Flt - Depress Man Weld To Continue FB1[301].22'; 9655 '~S001R08CN.I.Wc2SGunFlt - Weld Controller 2 Servo Gun Fault FB1[301].23'; 9656 '~S001R08CN.I.Wc2SGunMtrTempFlt - Cntrl 2 Servo Gun Motor Over Temp FB1[301].24'; 9657 '~S001R08CN.I.Td2MtrFlt - Tip Dress 2 Motor Fault FB1[301].25'; 9658 '~S001R08CN.I.WC2XfmrTempFlt - Weld Cntrl 2 Transformer Over Temp FB1[301].26'; 9659 '~S001R08CN.I.AutoTipChng2Flt - Auto Tip Changer 2 Fault FB1[301].27'; 9660 '~S001R08CN.I.Slr2NotReady - Seal Controller 2 Not Ready FB1[301].28'; 9661 '~S001R08CN.I.Slr2MajorFlt - Seal Controller 2 Major Fault FB1[301].29'; 9662 '~S001R08CN.I.Slr2VolNotOk - Seal Controller 2 Volume Not Ok Fault FB1[301].30'; 9663 '~S001R08CN.I.Slr2PurgeFlt - Seal Controller 2 Purge Fault FB1[301].31'; 9664 '~S001R08CN.I.Slr2DoserNot Filled - Seal Cntrl 2 Doser Not Filled FB1[302].0'; 9665 '~S001R08CN.I.Slr2No2ClnMxr - Seal Cntrl2 No 2C In Mixer Fault FB1[302].1'; 9666 '~S001R08CN.I.Slr2NzlBroken - Seal Controller 2 Nozzle Broken Fault FB1[302].2'; 9667 '~S001R08CN.I.Slr2NozzleChgReq - Seal Cntrl2 Nozzle Change Reqd FB1[302].3'; 9668 '~S001R08CN.I.Slr2CycleInterrupted - Seal Cntrl2 Cycle Interrupted FB1[302].4'; 9669 '~S001R08CN.I.Stdw2Flt - Stud Weld 2 Weld Fault FB1[302].5'; 9670 '~S001R08CN.I.Stdw2DlyExcdd - Stud Weld 2 Time Delay Exceeded Flt FB1[302].6'; 9671 '~S001R08CN.I.Stdw2Maint Reqd - Stud Weld 2 Maintenance Required FB1[302].7'; 9672 '~S001R08CN.I.Stdw2Reject - Stud Weld 2 art Reject Fault FB1[302].8'; 9673 '~S001R08CN.I.Rvt2Flt - Rivet Controller 2 Fault FB1[302].9'; 9674 '~S001R08CN.I.Rvt2DlyExcdd - Rivet Cntrl 2 Time Delay Exceeded Flt FB1[302].10'; 9675 '~S001R08CN.I.AutoPulledTipByp2 - Auto Pulled Tip Bypass 2 FB1[302].11'; 9676 '~S001R08CN.I.StdWld2EquipmentFlt - Stud Weld 2 Equipment Fault FB1[302].12'; 9677 '~S001R08CN.I.StdWld2BrcktNotPresent - Stud Weld 2 Bracket Not Pres FB1[302].13'; 9678 '~S001R08CN.Ix.LsrWldMntrFlt - Seam Geometry/Laser Weld Monitor Flt FB1[302].14'; 9679 '~S001R08CN.Ix.LsrHeadFlt - Laser Head Fault FB1[302].15'; 9680 '~S001R08CN.Ix.LsrGlsFlt - Glass Fault FB1[302].16'; 9681 '~S001R08CN.Ix.LsrWhlFlt - Pressure Wheel Not In Range Fault FB1[302].17'; 9682 '~S001R08CN.Ix.LsrGeoFlt - Seam Geometry/Laser Bad Process Geo Flt FB1[302].18'; 9683 '~S001R08CN.Ix.LsrHdCollFlt - Laser Head Collision Fault FB1[302].19'; 9684 '~S001R08CN.Ix.LsrHdSysFlt - Laser Head System Fault FB1[302].20'; 9685 '~S001R08CN.Ix.LsrHdFar - Laser Head Far Fault FB1[302].21'; 9686 '~S001R08CN.Ix.LsrHdSftCollFlt - Laser Head Software Collision Flt FB1[302].22'; 9687 '~S001R08CN.I.O.TipChngReqd2 - Weld Cntrl 2 Tip Change Required FB1[302].23'; 9688 '~S001R08CN.I.M.NutDetectFlt2 - Nut Welder 2 Nut Detection Fault FB1[302].24'; 9689 '~S001R08CN.I.M.NutProjFlt2 - Nut Welder 2 Weld Not In Tolerance FB1[302].25'; 9690 '~S001R08CN.I.TCWrongToolInStand - Tool Changer Wrong Tool In Stand FB1[302].26'; 9691 '~Spare FB1[302].27'; 9692 '~Spare FB1[302].28'; 9693 '~Spare FB1[302].29'; 9694 '~Spare FB1[302].30'; 9695 '~Spare FB1[302].31'; 9696 '~S001R08CN.I.VisionCommOK - Vision System Comm Fault FB1[303].0'; 9697 '~S001R08CN.I.OutOfTolerance - Vision System Out Of Tolerance FB1[303].1'; 9698 '~S001R08CN.I.MeasureReject - Vision System Measure Reject FB1[303].2'; 9699 '~S001R08CN.I.VisionSysCalibrationFlt - Vision System Calibration Flt FB1[303].3'; 9700 '~S001R08CN.I.VisionSysFlt - Vision System Flt FB1[303].4'; 9701 '~Spare FB1[303].5'; 9702 '~Spare FB1[303].6'; 9703 '~Spare FB1[303].7'; 9704 '~Spare FB1[303].8'; 9705 '~Spare FB1[303].9'; 9706 '~Spare FB1[303].10'; 9707 '~Spare FB1[303].11'; 9708 '~Spare FB1[303].12'; 9709 '~Spare FB1[303].13'; 9710 '~Spare FB1[303].14'; 9711 '~Spare FB1[303].15'; 9712 '~Spare FB1[303].16'; 9713 '~Spare FB1[303].17'; 9714 '~S001R08CN.M.InteruptCyc - Laser Cyc Interupt Cut Wire And Reject Car FB1[303].18'; 9715 '~S001R08CN.M.SuspectPart Inspect Vehicle And Accept Or Reject FB1[303].19'; 9716 '~S001R08 Power Meter High Power Fault Detected FB1[303].20'; 9717 '~S001R08 Power Meter Low Power Fault Detected FB1[303].21'; 9718 '~Spare FB1[303].22'; 9719 '~Spare FB1[303].23'; 9720 '~Spare FB1[303].24'; 9721 '~Spare FB1[303].25'; 9722 '~Spare FB1[303].26'; 9723 '~Spare FB1[303].27'; 9724 '~Spare FB1[303].28'; 9725 '~Spare FB1[303].29'; 9726 '~Spare FB1[303].30'; 9727 '~Spare FB1[303].31'; 9728 '~Spare FB1[304].0'; 9729 '~Spare FB1[304].1'; 9730 '~Spare FB1[304].2'; 9731 '~Spare FB1[304].3'; 9732 '~Spare FB1[304].4'; 9733 '~Spare FB1[304].5'; 9734 '~Spare FB1[304].6'; 9735 '~Spare FB1[304].7'; 9736 '~Spare FB1[304].8'; 9737 '~Spare FB1[304].9'; 9738 '~Spare FB1[304].10'; 9739 '~Spare FB1[304].11'; 9740 '~Spare FB1[304].12'; 9741 '~Spare FB1[304].13'; 9742 '~Spare FB1[304].14'; 9743 '~Spare FB1[304].15'; 9744 '~Spare FB1[304].16'; 9745 '~Spare FB1[304].17'; 9746 '~Spare FB1[304].18'; 9747 '~Spare FB1[304].19'; 9748 '~Spare FB1[304].20'; 9749 '~Spare FB1[304].21'; 9750 '~Spare FB1[304].22'; 9751 '~Spare FB1[304].23'; 9752 '~Spare FB1[304].24'; 9753 '~Spare FB1[304].25'; 9754 '~Spare FB1[304].26'; 9755 '~Spare FB1[304].27'; 9756 '~Spare FB1[304].28'; 9757 '~Spare FB1[304].29'; 9758 '~Spare FB1[304].30'; 9759 '~Spare FB1[304].31'; 9760 '~Spare FB1[305].0'; 9761 '~Spare FB1[305].1'; 9762 '~Spare FB1[305].2'; 9763 '~Spare FB1[305].3'; 9764 '~Spare FB1[305].4'; 9765 '~Spare FB1[305].5'; 9766 '~Spare FB1[305].6'; 9767 '~Spare FB1[305].7'; 9768 '~Spare FB1[305].8'; 9769 '~Spare FB1[305].9'; 9770 '~Spare FB1[305].10'; 9771 '~Spare FB1[305].11'; 9772 '~Spare FB1[305].12'; 9773 '~Spare FB1[305].13'; 9774 '~Spare FB1[305].14'; 9775 '~Spare FB1[305].15'; 9776 '~Spare FB1[305].16'; 9777 '~Spare FB1[305].17'; 9778 '~Spare FB1[305].18'; 9779 '~Spare FB1[305].19'; 9780 '~Spare FB1[305].20'; 9781 '~Spare FB1[305].21'; 9782 '~Spare FB1[305].22'; 9783 '~Spare FB1[305].23'; 9784 '~Spare FB1[305].24'; 9785 '~Spare FB1[305].25'; 9786 '~Spare FB1[305].26'; 9787 '~Spare FB1[305].27'; 9788 '~Spare FB1[305].28'; 9789 '~Spare FB1[305].29'; 9790 '~Spare FB1[305].30'; 9791 '~Spare FB1[305].31'; 9792 '~Spare FB1[306].0'; 9793 '~Spare FB1[306].1'; 9794 '~Spare FB1[306].2'; 9795 '~Spare FB1[306].3'; 9796 '~Spare FB1[306].4'; 9797 '~Spare FB1[306].5'; 9798 '~Spare FB1[306].6'; 9799 '~Spare FB1[306].7'; 9800 '~Spare FB1[306].8'; 9801 '~Spare FB1[306].9'; 9802 '~Spare FB1[306].10'; 9803 '~Spare FB1[306].11'; 9804 '~Spare FB1[306].12'; 9805 '~Spare FB1[306].13'; 9806 '~Spare FB1[306].14'; 9807 '~Spare FB1[306].15'; 9808 '~Spare FB1[306].16'; 9809 '~Spare FB1[306].17'; 9810 '~Spare FB1[306].18'; 9811 '~Spare FB1[306].19'; 9812 '~Spare FB1[306].20'; 9813 '~Spare FB1[306].21'; 9814 '~Spare FB1[306].22'; 9815 '~Spare FB1[306].23'; 9816 '~Spare FB1[306].24'; 9817 '~Spare FB1[306].25'; 9818 '~Spare FB1[306].26'; 9819 '~Spare FB1[306].27'; 9820 '~Spare FB1[306].28'; 9821 '~Spare FB1[306].29'; 9822 '~Spare FB1[306].30'; 9823 '~Spare FB1[306].31'; 9824 '~Spare FB1[307].0'; 9825 '~Spare FB1[307].1'; 9826 '~Spare FB1[307].2'; 9827 '~Spare FB1[307].3'; 9828 '~Spare FB1[307].4'; 9829 '~Spare FB1[307].5'; 9830 '~Spare FB1[307].6'; 9831 '~Spare FB1[307].7'; 9832 '~Spare FB1[307].8'; 9833 '~Spare FB1[307].9'; 9834 '~Spare FB1[307].10'; 9835 '~Spare FB1[307].11'; 9836 '~Spare FB1[307].12'; 9837 '~Spare FB1[307].13'; 9838 '~Spare FB1[307].14'; 9839 '~Spare FB1[307].15'; 9840 '~Spare FB1[307].16'; 9841 '~Spare FB1[307].17'; 9842 '~Spare FB1[307].18'; 9843 '~Spare FB1[307].19'; 9844 '~Spare FB1[307].20'; 9845 '~Spare FB1[307].21'; 9846 '~Spare FB1[307].22'; 9847 '~Spare FB1[307].23'; 9848 '~Spare FB1[307].24'; 9849 '~Spare FB1[307].25'; 9850 '~Spare FB1[307].26'; 9851 '~Spare FB1[307].27'; 9852 '~Spare FB1[307].28'; 9853 '~Spare FB1[307].29'; 9854 '~Spare FB1[307].30'; 9855 '~Spare FB1[307].31'; 9856 '~Spare FB1[308].0'; 9857 '~Spare FB1[308].1'; 9858 '~Spare FB1[308].2'; 9859 '~Spare FB1[308].3'; 9860 '~Spare FB1[308].4'; 9861 '~Spare FB1[308].5'; 9862 '~Spare FB1[308].6'; 9863 '~Spare FB1[308].7'; 9864 '~Spare FB1[308].8'; 9865 '~Spare FB1[308].9'; 9866 '~Spare FB1[308].10'; 9867 '~Spare FB1[308].11'; 9868 '~Spare FB1[308].12'; 9869 '~Spare FB1[308].13'; 9870 '~Spare FB1[308].14'; 9871 '~Spare FB1[308].15'; 9872 '~Spare FB1[308].16'; 9873 '~Spare FB1[308].17'; 9874 '~Spare FB1[308].18'; 9875 '~Spare FB1[308].19'; 9876 '~Spare FB1[308].20'; 9877 '~Spare FB1[308].21'; 9878 '~Spare FB1[308].22'; 9879 '~Spare FB1[308].23'; 9880 '~Spare FB1[308].24'; 9881 '~Spare FB1[308].25'; 9882 '~Spare FB1[308].26'; 9883 '~Spare FB1[308].27'; 9884 '~Spare FB1[308].28'; 9885 '~Spare FB1[308].29'; 9886 '~Spare FB1[308].30'; 9887 '~Spare FB1[308].31'; 9888 '~Spare FB1[309].0'; 9889 '~Spare FB1[309].1'; 9890 '~Spare FB1[309].2'; 9891 '~Spare FB1[309].3'; 9892 '~Spare FB1[309].4'; 9893 '~Spare FB1[309].5'; 9894 '~Spare FB1[309].6'; 9895 '~Spare FB1[309].7'; 9896 '~Spare FB1[309].8'; 9897 '~Spare FB1[309].9'; 9898 '~Spare FB1[309].10'; 9899 '~Spare FB1[309].11'; 9900 '~Spare FB1[309].12'; 9901 '~Spare FB1[309].13'; 9902 '~Spare FB1[309].14'; 9903 '~Spare FB1[309].15'; 9904 '~Spare FB1[309].16'; 9905 '~Spare FB1[309].17'; 9906 '~Spare FB1[309].18'; 9907 '~Spare FB1[309].19'; 9908 '~Spare FB1[309].20'; 9909 '~Spare FB1[309].21'; 9910 '~Spare FB1[309].22'; 9911 '~Spare FB1[309].23'; 9912 '~Spare FB1[309].24'; 9913 '~Spare FB1[309].25'; 9914 '~Spare FB1[309].26'; 9915 '~Spare FB1[309].27'; 9916 '~Spare FB1[309].28'; 9917 '~Spare FB1[309].29'; 9918 '~Spare FB1[309].30'; 9919 '~Spare FB1[309].31'; 9920 '~Spare FB1[310].0'; 9921 '~Spare FB1[310].1'; 9922 '~Spare FB1[310].2'; 9923 '~Spare FB1[310].3'; 9924 '~Spare FB1[310].4'; 9925 '~Spare FB1[310].5'; 9926 '~Spare FB1[310].6'; 9927 '~Spare FB1[310].7'; 9928 '~Spare FB1[310].8'; 9929 '~Spare FB1[310].9'; 9930 '~Spare FB1[310].10'; 9931 '~Spare FB1[310].11'; 9932 '~Spare FB1[310].12'; 9933 '~Spare FB1[310].13'; 9934 '~Spare FB1[310].14'; 9935 '~Spare FB1[310].15'; 9936 '~Spare FB1[310].16'; 9937 '~Spare FB1[310].17'; 9938 '~Spare FB1[310].18'; 9939 '~Spare FB1[310].19'; 9940 '~Spare FB1[310].20'; 9941 '~Spare FB1[310].21'; 9942 '~Spare FB1[310].22'; 9943 '~Spare FB1[310].23'; 9944 '~Spare FB1[310].24'; 9945 '~Spare FB1[310].25'; 9946 '~Spare FB1[310].26'; 9947 '~Spare FB1[310].27'; 9948 '~Spare FB1[310].28'; 9949 '~Spare FB1[310].29'; 9950 '~Spare FB1[310].30'; 9951 '~Spare FB1[310].31'; 9952 '~Spare FB1[311].0'; 9953 '~Spare FB1[311].1'; 9954 '~Spare FB1[311].2'; 9955 '~Spare FB1[311].3'; 9956 '~Spare FB1[311].4'; 9957 '~Spare FB1[311].5'; 9958 '~Spare FB1[311].6'; 9959 '~Spare FB1[311].7'; 9960 '~Spare FB1[311].8'; 9961 '~Spare FB1[311].9'; 9962 '~Spare FB1[311].10'; 9963 '~Spare FB1[311].11'; 9964 '~Spare FB1[311].12'; 9965 '~Spare FB1[311].13'; 9966 '~Spare FB1[311].14'; 9967 '~Spare FB1[311].15'; 9968 '~Spare FB1[311].16'; 9969 '~Spare FB1[311].17'; 9970 '~Spare FB1[311].18'; 9971 '~Spare FB1[311].19'; 9972 '~Spare FB1[311].20'; 9973 '~Spare FB1[311].21'; 9974 '~Spare FB1[311].22'; 9975 '~Spare FB1[311].23'; 9976 '~Spare FB1[311].24'; 9977 '~Spare FB1[311].25'; 9978 '~Spare FB1[311].26'; 9979 '~Spare FB1[311].27'; 9980 '~Spare FB1[311].28'; 9981 '~Spare FB1[311].29'; 9982 '~Spare FB1[311].30'; 9983 '~Spare FB1[311].31'; 9984 '~Spare FB1[312].0'; 9985 '~Spare FB1[312].1'; 9986 '~Spare FB1[312].2'; 9987 '~Spare FB1[312].3'; 9988 '~Spare FB1[312].4'; 9989 '~Spare FB1[312].5'; 9990 '~Spare FB1[312].6'; 9991 '~Spare FB1[312].7'; 9992 '~Spare FB1[312].8'; 9993 '~Spare FB1[312].9'; 9994 '~Spare FB1[312].10'; 9995 '~Spare FB1[312].11'; 9996 '~Spare FB1[312].12'; 9997 '~Spare FB1[312].13'; 9998 '~Spare FB1[312].14'; 9999 '~Spare FB1[312].15'; 10000 '**Local Message Display**'

text list "Text_list_IO_System": 1 'IO System 1'; 2 'IO System 2'; 3 'IO System 3'; 4 'IO System 4'

text list "G120D_Faults_Warnings": 1000 'F01000 - Internal software error'; 1001 'F01001 - FloatingPoint exception'; 1002 'F01002 - Internal software error'; 1003 'F01003 - Acknowledgment delay when accessing the memory'; 1004 'N01004 (F, A) - Internal software error'; 1005 'F01005 - File upload/download error'; 1009 'A01009 (N) - CU: Control module overtemperature'; 1010 'F01010 - Drive type unknown'; 1015 'F01015 - Internal software error'; 1016 'A01016 (F) - Firmware changed'; 1017 'A01017 - Component lists changed'; 1018 'F01018 - Booting has been interrupted several times'; 1019 'A01019 - Writing to the removable data medium unsuccessful'; 1020 'A01020 - Writing to RAM disk unsuccessful'; 1021 'A01021 - Removable data medium as USB data storage medium from the PC used'; 1023 'F01023 - Software timeout (internal)'; 1028 'A01028 (F) - Configuration error'; 1030 'F01030 - Sign-of-life failure for master control'; 1033 'F01033 - Units changeover: Reference parameter value invalid'; 1034 'F01034 - Units changeover: Calculation parameter values after reference value change unsuccessful'; 1035 'A01035 (F) - ACX: Parameter back-up file corrupted'; 1036 'F01036 (A) - ACX: Parameter back-up file missing'; 1038 'F01038 (A) - ACX: Loading the parameter back-up file unsuccessful'; 1039 'F01039 (A) - ACX: Writing to the parameter back-up file was unsuccessful'; 1040 'F01040 - Save parameter settings and carry out a POWER ON'; 1042 'F01042 - Parameter error during project download'; 1043 'F01043 - Fatal error at project download'; 1044 'F01044 - CU: Descriptive data error'; 1045 'A01045 - Configuring data invalid'; 1049 'A01049 - It is not possible to write to file'; 1054 'F01054 - CU: System limit exceeded'; 1064 'A01064 (F) - CU: Internal error (CRC)'; 1066 'A01066 - Buffer memory: 70% fill level reached or exceeded'; 1067 'A01067 - Buffer memory: 100 % fill level reached'; 1068 'F01068 - CU: Data memory memory overflow'; 1069 'A01069 - Parameter backup and device incompatible'; 1072 'F01072 - Memory card restored from the backup copy'; 1073 'A01073 (N) - POWER ON required for backup copy on memory card'; 1105 'F01105 (A) - CU: Insufficient memory'; 1107 'F01107 - Save to memory card unsuccessful'; 1112 'F01112 - CU: Power unit not permissible'; 1120 'F01120 (A) - Terminal initialization has failed'; 1122 'F01122 (A) - Frequency at the measuring probe input too high'; 1152 'F01152 - CU: Invalid constellation of drive object types'; 1205 'F01205 - CU: Time slice overflow'; 1250 'F01250 - CU: CU-EEPROM incorrect read-only data'; 1251 'A01251 - CU: CU-EEPROM incorrect read-write data'; 1257 'F01257 - CU: Firmware version out of date'; 1340 'F01340 - Topology: Too many components on one line'; 1505 'F01505 (A) - BICO: Interconnection cannot be established'; 1510 'F01510 - BICO: Signal source is not float type'; 1511 'F01511 (A) - BICO: Interconnection with different scalings'; 1512 'F01512 - BICO: No scaling available'; 1513 'F01513 (N, A) - BICO: Interconnection cross DO with different scalings'; 1514 'A01514 (F) - BICO: Error when writing during a reconnect'; 1515 'F01515 (A) - BICO: Writing to parameter not permitted as the master control is active'; 1590 'A01590 (F) - Drive: Motor maintenance interval expired'; 1600 'F01600 - SI P1 (CU): STOP A initiated'; 1611 'F01611 (A) - SI P1 (CU): Defect in a monitoring channel'; 1620 'N01620 (F, A) - SI P1 (CU): Safe Torque Off active'; 1625 'F01625 - SI P1 (CU): Sign-of-life error in safety data'; 1640 'F01640 - SI P1 (CU): component replacement identified and acknowledgment/save required'; 1641 'F01641 - SI P1 (CU): component replacement identified and save required'; 1649 'F01649 - SI P1 (CU): Internal software error'; 1650 'F01650 - SI P1 (CU): Acceptance test required'; 1651 'F01651 - SI P1 (CU): Synchronization safety time slices unsuccessful'; 1653 'F01653 - SI P1 (CU): PROFIBUS/PROFINET configuration error'; 1654 'A01654 (F) - SI P1 (CU): Deviating PROFIsafe configuration'; 1655 'F01655 - SI P1 (CU): Align monitoring functions'; 1656 'F01656 - SI P1 (CU): Parameter processor 2 error'; 1658 'F01658 - SI P1 (CU): PROFIsafe telegram number not suitable'; 1659 'F01659 - SI P1 (CU): Write request for parameter rejected'; 1660 'F01660 - SI P1 (CU): Safety-related functions not supported'; 1661 'F01661 - SI P1 (CU): Simulation of the safety inputs active'; 1662 'F01662 - Error internal communications'; 1663 'F01663 - SI P1 (CU): Copying the SI parameters rejected'; 1665 'F01665 - SI P1 (CU): System is defective'; 1666 'A01666 (F) - SI Motion P1 (CU): Steady-state (static) 1 signal at the F-DI for safe acknowledgment'; 1669 'A01669 (F, N) - SI Motion: Unfavorable combination of motor and power unit'; 1680 'F01680 - SI Motion P1 (CU): Checksum error safety monitoring functions'; 1681 'F01681 - SI Motion P1 (CU): Incorrect parameter value'; 1682 'F01682 - SI Motion P1 (CU): Monitoring function not supported'; 1683 'F01683 - SI Motion P1 (CU): SLS enable missing'; 1690 'F01690 - SI Motion: Data save problem for the NVRAM'; 1692 'F01692 - SI Motion P1 (CU): Parameter value not permitted for encoderless'; 1693 'A01693 (F) - SI P1 (CU): Safety parameter setting changed, POWER ON required'; 1696 'A01696 (F) - SI Motion: Test stop for the motion monitoring functions selected when booting'; 1697 'A01697 (F) - SI Motion: Test stop for motion monitoring functions required'; 1698 'A01698 (F) - SI P1 (CU): Commissioning mode active'; 1699 'A01699 (F) - SI P1 (CU): Test stop for STO required'; 1700 'C01700 - SI Motion P1 (CU): STOP A initiated'; 1701 'C01701 - SI Motion P1 (CU): STOP B initiated'; 1706 'C01706 - SI Motion P1 (CU): SAM/SBR limit exceeded'; 1711 'C01711 - SI Motion P1 (CU): Defect in a monitoring channel'; 1712 'C01712 - SI Motion P1 (CU): Defect in F-IO processing'; 1714 'C01714 - SI Motion P1 (CU): Safely Limited Speed exceeded'; 1716 'C01716 - SI Motion P1 (CU): Tolerance for safe motion direction exceeded'; 1770 'C01770 - SI Motion P1 (CU): Discrepancy error of the fail-safe inputs'; 1772 'A01772 - SI Motion P1 (CU): Test stop for fail-safe digital outputs running'; 1773 'F01773 - SI Motion P1 (CU): Test stop fail-safe digital output error'; 1774 'A01774 - SI Motion P1 (CU): Test stop for fail-safe digital outputs required'; 1788 'A01788 - SI: Automatic test stop waits for STO deselection via motion monitoring functions'; 1790 'A01790 - SI: Power up stopped due to STO via terminals'; 1796 'A01796 (F, N) - SI P1 (CU): Wait for communication'; 1798 'C01798 - SI Motion P1 (CU): Test stop for motion monitoring functions running'; 1799 'C01799 - SI Motion P1 (CU): Acceptance test mode active'; 1900 'A01900 (F) - PROFIBUS: Configuration telegram error'; 1910 'F01910 (N, A) - Fieldbus interface setpoint timeout'; 1920 'A01920 (F) - PROFIBUS: Interruption cyclic connection'; 1945 'A01945 - PROFIBUS: Connection to the Publisher failed'; 1946 'F01946 (A) - PROFIBUS: Connection to the Publisher aborted'; 1951 'F01951 - CU SYNC: Synchronization application clock cycle missing'; 1953 'A01953 - CU SYNC: Synchronization not completed'; 2050 'A02050 - Trace: Start not possible'; 2051 'A02051 - Trace: recording not possible as a result of know-how protection'; 2055 'A02055 - Trace: Recording time too short'; 2056 'A02056 - Trace: Recording cycle too short'; 2057 'A02057 - Trace: Time slice clock cycle invalid'; 2058 'A02058 - Trace: Time slice clock cycle for endless trace not valid'; 2059 'A02059 - Trace: Time slice clock cycle for 2 x 8 recording channels not valid'; 2060 'A02060 - Trace: Signal to be traced missing'; 2061 'A02061 - Trace: Invalid signal'; 2062 'A02062 - Trace: Invalid trigger signal'; 2063 'A02063 - Trace: Invalid data type'; 2070 'A02070 - Trace: Parameter cannot be changed'; 2075 'A02075 - Trace: Pretrigger time too long'; 2080 'F02080 - Trace: Parameterization deleted due to unit changeover'; 2095 'A02095 - MTrace 0: multiple trace cannot be activated'; 2096 'A02096 - MTrace 0: cannot be saved'; 2097 'A02097 - MTrace 1: multiple trace cannot be activated'; 2098 'A02098 - MTrace 1: cannot be saved'; 2099 'A02099 - Trace: Insufficient Control Unit memory'; 2150 'A02150 - OA: Application cannot be loaded'; 2151 'F02151 (A) - OA: Internal software error'; 2152 'F02152 (A) - OA: Insufficient memory'; 3000 'F03000 - NVRAM fault on action'; 3001 'F03001 - NVRAM checksum incorrect'; 3505 'F03505 (N, A) - Analog input wire breakage'; 3510 'A03510 (F, N) - Calibration data not plausible'; 5000 'A05000 (N) - Power unit: Overtemperature heat sink AC inverter'; 5001 'A05001 (N) - Power unit: Overtemperature depletion layer chip'; 5002 'A05002 (N) - Power unit: Air intake overtemperature'; 5004 'A05004 (N) - Power unit: Rectifier overtemperature'; 5006 'A05006 (N) - Power unit: Overtemperature thermal model'; 5065 'A05065 (F, N) - Voltage measured values not plausible'; 6310 'F06310 (A) - Supply voltage (p0210) incorrectly parameterized'; 6921 'A06921 (N) - Braking resistor phase unsymmetry'; 6922 'F06922 - Braking resistor phase failure'; 7011 'F07011 - Drive: Motor overtemperature'; 7012 'A07012 (N) - Drive: Motor temperature model 1/3 overtemperature'; 7014 'A07014 (N) - Drive: Motor temperature model configuration alarm'; 7015 'A07015 - Drive: Motor temperature sensor alarm'; 7016 'F07016 - Drive: Motor temperature sensor fault'; 7080 'F07080 - Drive: Incorrect control parameter'; 7082 'F07082 - Macro: Execution not possible'; 7083 'F07083 - Macro: ACX file not found'; 7084 'F07084 - Macro: Condition for WaitUntil not fulfilled'; 7086 'F07086 - Units changeover: Parameter limit violation due to reference value change'; 7088 'F07088 - Units changeover: Parameter limit violation due to units changeover'; 7089 'A07089 - Changing over units: Function module activation is blocked because the units have been changed over'; 7092 'A07092 - Drive: moment of inertia estimator still not ready'; 7094 'A07094 - General parameter limit violation'; 7200 'A07200 - Drive: Master control ON command present'; 7220 'F07220 (N, A) - Drive: Master control by PLC missing'; 7300 'F07300 (A) - Drive: Line contactor feedback signal missing'; 7320 'F07320 - Drive: Automatic restart interrupted'; 7321 'A07321 - Drive: Automatic restart active'; 7330 'F07330 - Flying restart: Measured search current too low'; 7331 'F07331 - Flying restart: Function not supported'; 7404 'F07404 - Drive: DC link voltage monitoring Vdc_max'; 7409 'A07409 (N) - Drive: U/f control, current limiting controller active'; 7410 'F07410 - Drive: Current controller output limited'; 7411 'F07411 - Drive: Flux setpoint not reached when building up excitation'; 7416 'A07416 - Drive: Flux controller configuration'; 7426 'F07426 (A) - Technology controller actual value limited'; 7428 'A07428 (N) - Technology controller parameterizing error'; 7435 'F07435 (N) - Drive: Setting the ramp-function generator for sensorless vector control'; 7440 'A07440 - EPOS: Jerk time is limited'; 7441 'A07441 - LR: Save the position offset of the absolute encoder adjustment'; 7442 'F07442 (A) - LR: Multiturn does not match the modulo range'; 7443 'F07443 (A) - LR: Reference point coordinate not in the permissible range'; 7450 'F07450 (A) - LR: Standstill monitoring has responded'; 7451 'F07451 (A) - LR: Position monitoring has responded'; 7452 'F07452 (A) - LR: Following error too high'; 7453 'F07453 - LR: Position actual value preprocessing error'; 7454 'A07454 - LR: Position actual value preprocessing does not have a valid encoder'; 7455 'A07455 - EPOS: Maximum velocity limited'; 7456 'A07456 - EPOS: Setpoint velocity limited'; 7457 'A07457 - EPOS: Combination of input signals illegal'; 7458 'F07458 - EPOS: Reference cam not found'; 7459 'F07459 - EPOS: No zero mark'; 7460 'F07460 - EPOS: End of reference cam not found'; 7461 'A07461 - EPOS: Reference point not set'; 7462 'A07462 - EPOS: Selected traversing block number does not exist'; 7463 'A07463 (F) - EPOS: External block change not requested in the traversing block'; 7464 'F07464 - EPOS: Traversing block is inconsistent'; 7465 'A07465 - EPOS: Traversing block does not have a subsequent block'; 7466 'A07466 - EPOS: Traversing block number assigned a multiple number of times'; 7467 'A07467 - EPOS: Traversing block has illegal task parameters'; 7468 'A07468 - EPOS: Traversing block jump destination does not exist'; 7469 'A07469 - EPOS: Traversing block < target position < software limit switch minus'; 7470 'A07470 - EPOS: Traversing block> target position > software limit switch plus'; 7471 'A07471 - EPOS: Traversing block target position outside the modulo range'; 7472 'A07472 - EPOS: Traversing block ABS_POS/ABS_NEG not possible'; 7473 'A07473 (F) - EPOS: Beginning of traversing range reached'; 7474 'A07474 (F) - EPOS: End of traversing range reached'; 7475 'F07475 (A) - EPOS: Target position < start of traversing range'; 7476 'F07476 (A) - EPOS: Target position > end of the traversing range'; 7477 'A07477 (F) - EPOS: Target position < software limit switch minus'; 7478 'A07478 (F) - EPOS: Target position > software limit switch plus'; 7479 'A07479 - EPOS: Software limit switch minus reached'; 7480 'A07480 - EPOS: Software limit switch plus reached'; 7481 'F07481 (A) - EPOS: Axis position < software limit switch minus'; 7482 'F07482 (A) - EPOS: Axis position > software limit switch plus'; 7483 'A07483 - EPOS: Travel to fixed stop clamping torque not reached'; 7484 'F07484 - EPOS: Fixed stop outside the monitoring window'; 7485 'F07485 (A) - EPOS: Fixed stop not reached'; 7486 'A07486 - EPOS: Intermediate stop missing'; 7487 'A07487 - EPOS: Reject traversing task missing'; 7488 'F07488 - EPOS: Relative positioning not possible'; 7489 'A07489 - EPOS: Reference point correction outside the window'; 7490 'F07490 (N) - EPOS: Enable signal withdrawn while traversing'; 7491 'F07491 (A) - EPOS: STOP cam minus reached'; 7492 'F07492 (A) - EPOS: STOP cam plus reached'; 7493 'F07493 - LR: Overflow of the value range for position actual value'; 7494 'F07494 - LR: Drive Data Set changeover in operation'; 7495 'A07495 (F) - LR: Reference function interrupted'; 7496 'A07496 - EPOS: Enable not possible'; 7497 'A07497 (N) - LR: Position setting value activated'; 7498 'A07498 (F) - LR: Measuring probe evaluation not possible'; 7499 'F07499 (A) - EPOS: Reversing cam approached with the incorrect traversing direction'; 7503 'F07503 - EPOS: STOP cam approached with the incorrect traversing direction'; 7505 'A07505 - EPOS: Task fixed stop not possible in the U/f/SLVC mode'; 7530 'A07530 - Drive: Drive Data Set DDS not present'; 7531 'A07531 - Drive: Command Data Set CDS not present'; 7550 'A07550 (F, N) - Drive: Not possible to reset encoder parameters'; 7552 'F07552 (A) - Drive encoder: Encoder configuration not supported'; 7553 'F07553 (A) - Drive encoder: Sensor Module configuration not supported'; 7557 'A07557 (F) - Encoder 1: Reference point coordinate not in the permissible range'; 7558 'A07558 (F) - Encoder 2: Reference point coordinate not in the permissible range'; 7563 'F07563 (A) - Drive encoder: XIST1_ERW configuration incorrect'; 7565 'A07565 (F, N) - Drive: Encoder error in PROFIdrive encoder interface 1'; 7566 'A07566 (F, N) - Drive: Encoder error in PROFIdrive encoder interface 2'; 7569 'A07569 (F) - Enc identification active'; 7570 'N07570 (F) - Encoder identification data transfer running'; 7577 'A07577 (F) - Encoder 1: Measuring probe evaluation not possible'; 7578 'A07578 (F) - Encoder 2: Measuring probe evaluation not possible'; 7581 'A07581 (F) - Encoder 1: Position actual value preprocessing error'; 7582 'A07582 (F) - Encoder 2: Position actual value preprocessing error'; 7584 'A07584 - Encoder 1: Position setting value activated'; 7585 'A07585 - Encoder 2: Position setting value activated'; 7587 'A07587 - Encoder 1: Position actual value preprocessing does not have a valid encoder'; 7588 'A07588 - Encoder 2: Position actual value preprocessing does not have a valid encoder'; 7590 'A07590 (F) - Encoder 1: Drive Data Set changeover in operation'; 7591 'A07591 (F) - Encoder 2: Drive Data Set changeover in operation'; 7593 'A07593 (F, N) - Encoder 1: Value range for position actual value exceeded'; 7594 'A07594 (F, N) - Encoder 2: Value range for position actual value exceeded'; 7596 'A07596 (F) - Encoder 1: Reference function interrupted'; 7597 'A07597 (F) - Encoder 2: Reference function interrupted'; 7599 'F07599 (A) - Encoder 1: Adjustment not possible'; 7600 'F07600 (A) - Encoder 2: Adjustment not possible'; 7754 'F07754 - Drive: Incorrect shutoff valve configuration'; 7800 'F07800 - Drive: No power unit present'; 7801 'F07801 - Drive: Motor overcurrent'; 7802 'F07802 - Drive: Infeed or power unit not ready'; 7805 'A07805 (N) - Drive: Power unit overload I2t'; 7806 'F07806 - Drive: Regenerative power limit exceeded (F3E)'; 7807 'F07807 - Drive: Short-circuit/ground fault detected'; 7810 'F07810 - Drive: Power unit EEPROM without rated data'; 7850 'A07850 (F) - External alarm 1'; 7851 'A07851 (F) - External alarm 2'; 7852 'A07852 (F) - External alarm 3'; 7860 'F07860 (A) - External fault 1'; 7861 'F07861 (A) - External fault 2'; 7862 'F07862 (A) - External fault 3'; 7891 'A07891 - Drive: Load monitoring pump/fan blocked'; 7892 'A07892 - Drive: Load monitoring pump/fan no load condition'; 7893 'A07893 - Drive: Load monitoring pump leakage'; 7894 'F07894 - Drive: Load monitoring pump/fan blocked'; 7895 'F07895 - Drive: Load monitoring pump/fan no load condition'; 7896 'F07896 - Drive: Load monitoring pump leakage'; 7900 'F07900 (N, A) - Drive: Motor blocked'; 7901 'F07901 - Drive: Motor overspeed'; 7902 'F07902 (N, A) - Drive: Motor stalled'; 7903 'A07903 - Drive: Motor speed deviation'; 7910 'A07910 (N) - Drive: Motor overtemperature'; 7920 'A07920 - Drive: Torque/speed too low'; 7921 'A07921 - Drive: Torque/speed too high'; 7922 'A07922 - Drive: Torque/speed out of tolerance'; 7923 'F07923 - Drive: Torque/speed too low'; 7924 'F07924 - Drive: Torque/speed too high'; 7925 'F07925 - Drive: Torque/speed out of tolerance'; 7926 'A07926 - Drive: Envelope curve parameter invalid'; 7927 'A07927 - DC braking active'; 7929 'A07929 (F) - Drive: No motor detected'; 7936 'F07936 - Drive: load failure'; 7950 'F07950 (A) - Motor parameter incorrect'; 7960 'A07960 - Drive: Incorrect friction characteristic'; 7961 'A07961 - Drive: Friction characteristic record activated'; 7963 'F07963 - Drive: Friction characteristic record interrupted'; 7967 'F07967 - Drive: Incorrect pole position identification'; 7968 'F07968 - Drive: Lq-Ld measurement incorrect'; 7969 'F07969 - Drive: Incorrect pole position identification'; 7975 'A07975 (N) - Drive: Travel to the zero mark - setpoint input expected'; 7980 'A07980 - Drive: Rotating measurement activated'; 7981 'A07981 - Drive: Enable signals for the rotating measurement missing'; 7982 'F07982 - Drive: Rotating measurement encoder test'; 7983 'F07983 - Drive: Rotating measurement saturation characteristic'; 7984 'F07984 - Drive: Speed controller optimization, moment of inertia'; 7985 'F07985 - Drive: Speed controller optimization (oscillation test)'; 7986 'F07986 - Drive: Rotating measurement ramp-function generator'; 7988 'F07988 - Drive: Rotating measurement, no configuration selected'; 7990 'F07990 - Drive: Incorrect motor data identification'; 7991 'A07991 (N) - Drive: Motor data identification activated'; 7994 'A07994 (F, N) - Drive: motor data identification not performed'; 8010 'F08010 (N, A) - CU: Analog-to-digital converter'; 8501 'F08501 (N, A) - PROFINET: Setpoint timeout'; 8502 'F08502 (A) - PROFINET: Monitoring time sign-of-life expired'; 8511 'A08511 (F) - PROFINET: Receive configuration data invalid'; 8526 'A08526 (F) - PROFINET: No cyclic connection'; 8564 'A08564 - PN/COMM BOARD: syntax error in the configuration file'; 8565 'A08565 - PROFINET: Consistency error affecting adjustable parameters'; 8760 'A08760 - CAN: maximum size of the IF PZD exceeded'; 8800 'A08800 